// TIA Portal project "XSFW_TIA60401_A3_V14_V15.1" (V15.1) (continued)
   "AuxTempMS050" AT %MW340 : Int;
   "AuxTempMS051" AT %MW342 : Int;
   "AuxTempMS052" AT %MW344 : Int;
   "AuxTempMS053" AT %MW346 : Int;
   "AuxTempMS054" AT %MW348 : Int;
   "AuxTempMS055" AT %MW350 : Int;
   "AuxTempMS056" AT %MW352 : Int;
   "AuxTempMC060" AT %MW354 : Int;
   "AuxTempMC061" AT %MW356 : Int;
   "AuxTempMC062" AT %MW358 : Int;
   "AuxTempMC063" AT %MW360 : Int;
   "AuxTempMC064" AT %MW362 : Int;
   "AuxTempMC065" AT %MW364 : Int;
   "ProxMantBoost1" AT %MD16 : DInt;
   "LimiteMantBoost1" AT %M1.7 : Bool;
   "ProxMantBoost2" AT %MD26 : DInt;
   "LimiteMantBoost2" AT %M2.3 : Bool;
END_VAR

DATA_BLOCK "DB_Fecha"   // DB1
{ S7_Optimized_Access := 'FALSE' }
VERSION : 0.1
   VAR
      STAT0 : Date_And_Time := DT#12-7-5-15:25:53.162;
      STAT1 : Int := 15;
      STAT2 : Int := 25;
      STAT3 : Int := 53;
      STAT4 : Int := 5;
      STAT5 : Int := 7;
      STAT6 : Int := 15;
      STAT7 : Int := 18;
      STAT8 : Int;
      STAT9 : Int := 8;
      STAT10 : Int;
      STAT11 : Word := W#16#15;
      STAT12 : Word := W#16#25;
      STAT13 : Word := W#16#53;
      STAT14 : Word := W#16#5;
      STAT15 : Word := W#16#7;
      STAT16 : Word := W#16#12;
   END_VAR
BEGIN
END_DATA_BLOCK

DATA_BLOCK "Enclavamientos"   // DB28
{ S7_Optimized_Access := 'FALSE' }
VERSION : 0.1
   VAR
      En1 : Bool := true;
      En2 : Bool := true;
      En3 : Bool;
      En4 : Bool;
      En5 : Bool;
      En6 : Bool;
      En7 : Bool;
      En8 : Bool;
      En9 : Bool;
      En10 : Bool;
      En11 : Bool;
      En12 : Bool;
      En13 : Bool;
      En14 : Bool;
      En15 : Bool;
      En16 : Bool;
      En17 : Bool;
      En18 : Bool;
      En19 : Bool;
      En20 : Bool;
      En21 : Bool;
      En22 : Bool;
      En23 : Bool;
      En24 : Bool;
      En25 : Bool;
      En26 : Bool;
      En27 : Bool;
      En28 : Bool;
      En29 : Bool;
      En30 : Bool;
      En31 : Bool;
      En32 : Bool;
      En33 : Bool;
      En34 : Bool;
      En35 : Bool;
      En36 : Bool;
      En37 : Bool;
      En38 : Bool;
      En39 : Bool;
      En40 : Bool;
      En41 : Bool;
      En42 : Bool;
      En43 : Bool;
      En44 : Bool;
      En45 : Bool;
      En46 : Bool;
      En47 : Bool;
      En48 : Bool;
      En49 : Bool;
      En50 : Bool;
      En51 : Bool;
      En52 : Bool;
      En53 : Bool;
      En54 : Bool;
      En55 : Bool;
      En56 : Bool;
      En57 : Bool;
      En58 : Bool;
      En59 : Bool;
      En60 : Bool;
      En61 : Bool;
      En62 : Bool;
      En63 : Bool;
      En64 : Bool;
   END_VAR
BEGIN
END_DATA_BLOCK

// folder: Alarmas

DATA_BLOCK "DB_ALA_PRE"   // DB32
{ S7_Optimized_Access := 'FALSE' }
VERSION : 0.1
   VAR
      x : Bool;   // Ninguna bomba de intercambiador de soplado en marcha
      x1 : Bool;   // Ninguna bomba de chillers de soplado en marcha
      x2 : Bool;   // Ninguna bomba de intercambiador de envasado en marcha
      x3 : Bool;   // Ninguna bomba de chillers de envasado en marcha
      x4 : Bool;   // Ninguna bomba de torre de enfiamiento de chillers en marcha
      x5 : Bool;   // Ningún Chiller de soplado habilitado
      x6 : Bool;   // Ningún chiller de envasado habilitado
      x7 : Bool;   // Alarma Presente en Chiller de soplado Grande
      x8 : Bool;   // Alarma Presente en Chiller de envasado Grande
      x9 : Bool;   // Chiller de soplado Grande en su máxima capacidad
      x10 : Bool;   // Chiller de envasado Grande en su máxima capacidad
      x11 : Bool;   // Falla Térmico MT007
      x12 : Bool;   // Falla Contactor MT007
      x13 : Bool;   // Falla Térmico MT008
      x14 : Bool;   // Falla Contactor MT008
      x15 : Bool;   // Falla Térmico MT009
      x16 : Bool;   // Falla Contactor MT009
      x17 : Bool;   // Falla Térmico MT010
      x18 : Bool;   // Falla Contactor MT010
      x19 : Bool;   // Falla Térmico MP010
      x20 : Bool;   // Falla Contactor MP010
      x21 : Bool;   // Falla Térmico MP011
      x22 : Bool;   // Falla Contactor MP011
      x23 : Bool;   // Falla Térmico MP012
      x24 : Bool;   // Falla Contactor MP012
      x25 : Bool;   // Falla Térmico MP013
      x26 : Bool;   // Falla Contactor MP013
      x27 : Bool;   // Falla Térmico MP018
      x28 : Bool;   // Falla Contactor MP018
      x29 : Bool;   // Falla Térmico MP019
      x30 : Bool;   // Falla Contactor MP019
      x31 : Bool;   // Falla Térmico V001
      x32 : Bool;   // Falla Contactor V001
      x33 : Bool;   // Falla Térmico V002
      x34 : Bool;   // Falla Contactor V002
      x35 : Bool;   // Falla Térmico V003
      x36 : Bool;   // Falla Contactor V003
      x37 : Bool;   // Falla Térmico MC060
      x38 : Bool;   // Falla Contactor MC060
      x39 : Bool;   // Falla Térmico MC061
      x40 : Bool;   // Falla Contactor MC061
      x41 : Bool;   // Falla Térmico MC062
      x42 : Bool;   // Falla Contactor MC062
      x43 : Bool;   // Falla Térmico MC063
      x44 : Bool;   // Falla Contactor MC063
      x45 : Bool;   // Falla Térmico MC064
      x46 : Bool;   // Falla Contactor MC064
      x47 : Bool;   // Falla Térmico MS050
      x48 : Bool;   // Falla Contactor MS050
      x49 : Bool;   // Falla Térmico MS051
      x50 : Bool;   // Falla Contactor MS051
      x51 : Bool;   // Falla Térmico MS052
      x52 : Bool;   // Falla Contactor MS052
      x53 : Bool;   // Falla Térmico MS053
      x54 : Bool;   // Falla Contactor MS053
      x55 : Bool;   // Falla Presostato Chillers
      x56 : Bool;   // Falla Térmico MS054
      x57 : Bool;   // Falla Contactor MS054
      x58 : Bool;   // Falla Térmico MS055
      x59 : Bool;   // Falla Contactor MS055
      x60 : Bool;   // Falla Térmico MV030
      x61 : Bool;   // Falla Contactor MV030
      x62 : Bool;   // Falla Térmico MV031
      x63 : Bool;   // Falla Contactor MV031
      x64 : Bool;   // Falla Térmico MP014
      x65 : Bool;   // Falla Contactor MP014
      x66 : Bool;   // Falla Térmico MP015
      x67 : Bool;   // Falla Contactor MP015
      x68 : Bool;   // Falla Térmico MC001
      x69 : Bool;   // Falla Contactor MC001
      x70 : Bool;   // Falla Térmico MC002
      x71 : Bool;   // Falla Contactor MC002
      x72 : Bool;   // Falla Térmico MC003
      x73 : Bool;   // Falla Contactor MC003
      x74 : Bool;   // Falla Térmico MC004
      x75 : Bool;   // Falla Contactor MC004
      x76 : Bool;   // Falla Térmico MC005
      x77 : Bool;   // Falla Contactor MC005
      x78 : Bool;   // Falla Flujostato Torres Cavaleto
      x79 : Bool;   // Falla Compresor ABC2 Baja Presion de Aceite
      x80 : Bool;   // Falla Compresor ABC2 Baja Presion de Agua
      x81 : Bool;   // Falla Compresor ABC2 Alta Temperatura de Aire
      x82 : Bool;   // Falla Compresor ABC2 Alta Temperatura de agua
      x83 : Bool;   // Falla Compresor ABC3 Baja Presion de Aceite
      x84 : Bool;   // Falla Compresor ABC3 Baja Presion de Agua
      x85 : Bool;   // Falla Compresor ABC3 Alta Temperatura de Aire
      x86 : Bool;   // Falla Compresor ABC3 Alta Temperatura de agua
      x87 : Bool;   // Falla Compresor ABC4 Baja Presion de Aceite
      x88 : Bool;   // Falla Compresor ABC4 Alta Temperatura de Aire
      x89 : Bool;   // Falla Compresor ABC4 Alta Temperatura de Aire
      x90 : Bool;   // Falla Compresor ABC4 Alta Temperatura de agua
      x91 : Bool;   // Falla Compresor ABC5 Baja Presion de Aceite
      x92 : Bool;   // Falla Compresor ABC5 Alta Temperatura de Aire
      x93 : Bool;   // Falla Compresor ABC5 Alta Temperatura de Aire
      x94 : Bool;   // Falla Compresor ABC5 Alta Temperatura de agua
      x95 : Bool;   // Falla Compresor Bellis & MHW28 Baja Presion Aceite
      x96 : Bool;   // Falla Compresor Bellis & MHW28 Baja Presion de Agua
      x97 : Bool;   // Falla Compresor Bellis & MHW28 Alta temperatura de Aire
      x98 : Bool;   // Falla Compresor Bellis & MHW28 Alta temperatura de Agua
      x99 : Bool;   // Falla Compresor Bellis & MHW28 Falla de Flujostato
      x100 : Bool;   // Requiere Marcha MC001
      x101 : Bool;   // Requiere Marcha MC002
      x102 : Bool;   // Requiere Marcha MC003
      x103 : Bool;   // Requiere Marcha MC004
      x104 : Bool;   // Requiere Marcha MC005
      x105 : Bool;   // Falla Conexión con sensor de Temperatura torres de Cavaleto
      x106 : Bool;   // Falla Conexión con sensor de Temperatura torres de Chillers
      x107 : Bool;   // Falla Conexión con sensor de Presión de ALTA
      x108 : Bool;   // Falla Conexión con sensor de Presión de ALTA redundante
      x109 : Bool;   // Falla Conexión con sensor de Presión de Baja
      x110 : Bool;   // Falla Presión de Alta en Límite Mínimo
      x111 : Bool;   // Falla Presión de Alta en demasiado Baja
      x112 : Bool;   // Falla Presión de Alta en demasiado Alta
      x113 : Bool;   // Falla Presión de Alta en Límite Máximo
      x114 : Bool;   // Falla Presión de Baja en Límite Mínimo
      x115 : Bool;   // Falla Presión de Baja en demasiado Baja
      x116 : Bool;   // Falla Presión de Baja en demasiado Alta
      x117 : Bool;   // Falla Presión de Baja en Límite Máximo
      x118 : Bool;   // Falla en chiller de envasado chico
      x119 : Bool;   // Falla en chiller de soplado chico
      x120 : Bool;   // Horas máximas en Compresor 1
      x121 : Bool;   // Horas máximas en Compresor 2
      x122 : Bool;   // Horas máximas en Compresor 3
      x123 : Bool;   // Horas máximas en Compresor 4
      x124 : Bool;   // Horas máximas en Compresor 5
      x125 : Bool;   // Falla algún contactor en Booster
      x126 : Bool;   // Falla algún guardamotor en Booster
      x127 : Bool;   // Presión Alta en Booster
      x128 : Bool;   // Falla algún contactor en Booster 2
      x129 : Bool;   // Falla algún guardamotor en Booster 2
      x130 : Bool;   // Error lectura analógica Presión Boosters
      x131 : Bool;   // Libre
      x132 : Bool;   // Libre
      x133 : Bool;   // Libre
      x134 : Bool;   // Libre
      x135 : Bool;   // Libre
      x136 : Bool;   // Libre
      x137 : Bool;   // Libre
      x138 : Bool;   // Libre
      x139 : Bool;   // Libre
      x140 : Bool;   // Libre
      x141 : Bool;   // Libre
      x142 : Bool;   // Libre
      x143 : Bool;   // Libre
      x144 : Bool;   // ABC1 TTA
      x145 : Bool;   // ABC1TTB
      x146 : Bool;   // ABC1PTA
      x147 : Bool;   // ABC1PTB
      x148 : Bool;   // ABC1Termico
      x149 : Bool;   // ABC1Confirmacion
      x150 : Bool;
      x151 : Bool;
      x152 : Bool;
      x153 : Bool;
      x154 : Bool;
      x155 : Bool;
      x156 : Bool;
      x157 : Bool;
      x158 : Bool;
      x159 : Bool;
      x160 : Bool;
      x161 : Bool;
      x162 : Bool;
      x163 : Bool;
      x164 : Bool;
      x165 : Bool;
      x166 : Bool;
      x167 : Bool;
      x168 : Bool;
      x169 : Bool;
      x170 : Bool;
      x171 : Bool;
      x172 : Bool;
      x173 : Bool;
      x174 : Bool;
      x175 : Bool;
      x176 : Bool;
      x177 : Bool;
      x178 : Bool;
      x179 : Bool;
      x180 : Bool;
      x181 : Bool;
      x182 : Bool;
      x183 : Bool;
      x184 : Bool;
      x185 : Bool;
      x186 : Bool;
      x187 : Bool;
      x188 : Bool;
      x189 : Bool;
      x190 : Bool;
      x191 : Bool;
      x192 : Bool;
      x193 : Bool;
      x194 : Bool;
      x195 : Bool;
      x196 : Bool;
      x197 : Bool;
      x198 : Bool;
      x199 : Bool;
   END_VAR
BEGIN
END_DATA_BLOCK

DATA_BLOCK "DB_ALA_REC"   // DB33
{ S7_Optimized_Access := 'FALSE' }
VERSION : 0.1
   VAR
      x : Bool;   // Ninguna bomba de intercambiador de soplado en marcha
      x1 : Bool;   // Ninguna bomba de chillers de soplado en marcha
      x2 : Bool;   // Ninguna bomba de intercambiador de envasado en marcha
      x3 : Bool;   // Ninguna bomba de chillers de envasado en marcha
      x4 : Bool;   // Ninguna bomba de torre de enfiamiento de chillers en marcha
      x5 : Bool;   // Ningún Chiller de soplado habilitado
      x6 : Bool;   // Ningún chiller de envasado habilitado
      x7 : Bool;   // Alarma Presente en Chiller de soplado Grande
      x8 : Bool;   // Alarma Presente en Chiller de envasado Grande
      x9 : Bool;   // Chiller de soplado Grande en su máxima capacidad
      x10 : Bool;   // Chiller de envasado Grande en su máxima capacidad
      x11 : Bool;   // Falla Térmico MT007
      x12 : Bool;   // Falla Contactor MT007
      x13 : Bool;   // Falla Térmico MT008
      x14 : Bool;   // Falla Contactor MT008
      x15 : Bool;   // Falla Térmico MT009
      x16 : Bool;   // Falla Contactor MT009
      x17 : Bool;   // Falla Térmico MT010
      x18 : Bool;   // Falla Contactor MT010
      x19 : Bool;   // Falla Térmico MP010
      x20 : Bool;   // Falla Contactor MP010
      x21 : Bool;   // Falla Térmico MP011
      x22 : Bool;   // Falla Contactor MP011
      x23 : Bool;   // Falla Térmico MP012
      x24 : Bool;   // Falla Contactor MP012
      x25 : Bool;   // Falla Térmico MP013
      x26 : Bool;   // Falla Contactor MP013
      x27 : Bool;   // Falla Térmico MP018
      x28 : Bool;   // Falla Contactor MP018
      x29 : Bool;   // Falla Térmico MP019
      x30 : Bool;   // Falla Contactor MP019
      x31 : Bool;   // Falla Térmico V001
      x32 : Bool;   // Falla Contactor V001
      x33 : Bool;   // Falla Térmico V002
      x34 : Bool;   // Falla Contactor V002
      x35 : Bool;   // Falla Térmico V003
      x36 : Bool;   // Falla Contactor V003
      x37 : Bool;   // Falla Térmico MC060
      x38 : Bool;   // Falla Contactor MC060
      x39 : Bool;   // Falla Térmico MC061
      x40 : Bool;   // Falla Contactor MC061
      x41 : Bool;   // Falla Térmico MC062
      x42 : Bool;   // Falla Contactor MC062
      x43 : Bool;   // Falla Térmico MC063
      x44 : Bool;   // Falla Contactor MC063
      x45 : Bool;   // Falla Térmico MC064
      x46 : Bool;   // Falla Contactor MC064
      x47 : Bool;   // Falla Térmico MS050
      x48 : Bool;   // Falla Contactor MS050
      x49 : Bool;   // Falla Térmico MS051
      x50 : Bool;   // Falla Contactor MS051
      x51 : Bool;   // Falla Térmico MS052
      x52 : Bool;   // Falla Contactor MS052
      x53 : Bool;   // Falla Térmico MS053
      x54 : Bool;   // Falla Contactor MS053
      x55 : Bool;   // Falla Presostato Chillers
      x56 : Bool;   // Falla Térmico MS054
      x57 : Bool;   // Falla Contactor MS054
      x58 : Bool;   // Falla Térmico MS055
      x59 : Bool;   // Falla Contactor MS055
      x60 : Bool;   // Falla Térmico MV030
      x61 : Bool;   // Falla Contactor MV030
      x62 : Bool;   // Falla Térmico MV031
      x63 : Bool;   // Falla Contactor MV031
      x64 : Bool;   // Falla Térmico MP014
      x65 : Bool;   // Falla Contactor MP014
      x66 : Bool;   // Falla Térmico MP015
      x67 : Bool;   // Falla Contactor MP015
      x68 : Bool;   // Falla Térmico MC001
      x69 : Bool;   // Falla Contactor MC001
      x70 : Bool;   // Falla Térmico MC002
      x71 : Bool;   // Falla Contactor MC002
      x72 : Bool;   // Falla Térmico MC003
      x73 : Bool;   // Falla Contactor MC003
      x74 : Bool;   // Falla Térmico MC004
      x75 : Bool;   // Falla Contactor MC004
      x76 : Bool;   // Falla Térmico MC005
      x77 : Bool;   // Falla Contactor MC005
      x78 : Bool;   // Falla Flujostato Torres Cavaleto
      x79 : Bool;   // Falla Compresor ABC2 Baja Presion de Aceite
      x80 : Bool;   // Falla Compresor ABC2 Baja Presion de Agua
      x81 : Bool;   // Falla Compresor ABC2 Alta Temperatura de Aire
      x82 : Bool;   // Falla Compresor ABC2 Alta Temperatura de agua
      x83 : Bool;   // Falla Compresor ABC3 Baja Presion de Aceite
      x84 : Bool;   // Falla Compresor ABC3 Baja Presion de Agua
      x85 : Bool;   // Falla Compresor ABC3 Alta Temperatura de Aire
      x86 : Bool;   // Falla Compresor ABC3 Alta Temperatura de agua
      x87 : Bool;   // Falla Compresor ABC4 Baja Presion de Aceite
      x88 : Bool;   // Falla Compresor ABC4 Alta Temperatura de Aire
      x89 : Bool;   // Falla Compresor ABC4 Alta Temperatura de Aire
      x90 : Bool;   // Falla Compresor ABC4 Alta Temperatura de agua
      x91 : Bool;   // Falla Compresor ABC5 Baja Presion de Aceite
      x92 : Bool;   // Falla Compresor ABC5 Alta Temperatura de Aire
      x93 : Bool;   // Falla Compresor ABC5 Alta Temperatura de Aire
      x94 : Bool;   // Falla Compresor ABC5 Alta Temperatura de agua
      x95 : Bool;   // Falla Compresor Bellis & MHW28 Baja Presion Aceite
      x96 : Bool;   // Falla Compresor Bellis & MHW28 Baja Presion de Agua
      x97 : Bool;   // Falla Compresor Bellis & MHW28 Alta temperatura de Aire
      x98 : Bool;   // Falla Compresor Bellis & MHW28 Alta temperatura de Agua
      x99 : Bool;   // Falla Compresor Bellis & MHW28 Falla de Flujostato
      x100 : Bool;   // Requiere Marcha MC001
      x101 : Bool;   // Requiere Marcha MC002
      x102 : Bool;   // Requiere Marcha MC003
      x103 : Bool;   // Requiere Marcha MC004
      x104 : Bool;   // Requiere Marcha MC005
      x105 : Bool;   // Falla Conexión con sensor de Temperatura torres de Cavaleto
      x106 : Bool;   // Falla Conexión con sensor de Temperatura torres de Chillers
      x107 : Bool;   // Falla Conexión con sensor de Presión de ALTA
      x108 : Bool;   // Falla Conexión con sensor de Presión de ALTA redundante
      x109 : Bool;   // Falla Conexión con sensor de Presión de Baja
      x110 : Bool;   // Falla Presión de Alta en Límite Mínimo
      x111 : Bool;   // Falla Presión de Alta en demasiado Baja
      x112 : Bool;   // Falla Presión de Alta en demasiado Alta
      x113 : Bool;   // Falla Presión de Alta en Límite Máximo
      x114 : Bool;   // Falla Presión de Baja en Límite Mínimo
      x115 : Bool;   // Falla Presión de Baja en demasiado Baja
      x116 : Bool;   // Falla Presión de Baja en demasiado Alta
      x117 : Bool;   // Falla Presión de Baja en Límite Máximo
      x118 : Bool;   // Falla en chiller de envasado chico
      x119 : Bool;   // Falla en chiller de soplado chico
      x120 : Bool;   // Horas máximas en Compresor 1
      x121 : Bool;   // Horas máximas en Compresor 2
      x122 : Bool;   // Horas máximas en Compresor 3
      x123 : Bool;   // Horas máximas en Compresor 4
      x124 : Bool;   // Horas máximas en Compresor 5
      x125 : Bool;   // Falla algún contactor en Booster
      x126 : Bool;   // Falla algún guardamotor en Booster
      x127 : Bool;   // Presión Alta en Booster
      x128 : Bool;   // Falla algún contactor en Booster 2
      x129 : Bool;   // Falla algún guardamotor en Booster 2
      x130 : Bool;   // Error lectura analógica Presión Boosters
      x131 : Bool;   // Libre
      x132 : Bool;   // Libre
      x133 : Bool;   // Libre
      x134 : Bool;   // Libre
      x135 : Bool;   // Libre
      x136 : Bool;   // Libre
      x137 : Bool;   // Libre
      x138 : Bool;   // Libre
      x139 : Bool;   // Libre
      x140 : Bool;   // Libre
      x141 : Bool;   // Libre
      x142 : Bool;   // Libre
      x143 : Bool;   // Libre
      x144 : Bool;   // ABC1 TTA
      x145 : Bool;   // ABC1TTB
      x146 : Bool;   // ABC1PTA
      x147 : Bool;   // ABC1PTB
      x148 : Bool;   // ABC1Termico
      x149 : Bool;   // ABC1Confirmacion
      x150 : Bool;
      x151 : Bool;
      x152 : Bool;
      x153 : Bool;
      x154 : Bool;
      x155 : Bool;
      x156 : Bool;
      x157 : Bool;
      x158 : Bool;
      x159 : Bool;
      x160 : Bool;
      x161 : Bool;
      x162 : Bool;
      x163 : Bool;
      x164 : Bool;
      x165 : Bool;
      x166 : Bool;
      x167 : Bool;
      x168 : Bool;
      x169 : Bool;
      x170 : Bool;
      x171 : Bool;
      x172 : Bool;
      x173 : Bool;
      x174 : Bool;
      x175 : Bool;
      x176 : Bool;
      x177 : Bool;
      x178 : Bool;
      x179 : Bool;
      x180 : Bool;
      x181 : Bool;
      x182 : Bool;
      x183 : Bool;
      x184 : Bool;
      x185 : Bool;
      x186 : Bool;
      x187 : Bool;
      x188 : Bool;
      x189 : Bool;
      x190 : Bool;
      x191 : Bool;
      x192 : Bool;
      x193 : Bool;
      x194 : Bool;
      x195 : Bool;
      x196 : Bool;
      x197 : Bool;
      x198 : Bool;
      x199 : Bool;
   END_VAR
BEGIN
END_DATA_BLOCK

DATA_BLOCK "DB_ALA_MEM"   // DB34
{ S7_Optimized_Access := 'FALSE' }
VERSION : 0.1
   VAR
      x : Bool;   // Ninguna bomba de intercambiador de soplado en marcha
      x1 : Bool;   // Ninguna bomba de chillers de soplado en marcha
      x2 : Bool;   // Ninguna bomba de intercambiador de envasado en marcha
      x3 : Bool;   // Ninguna bomba de chillers de envasado en marcha
      x4 : Bool;   // Ninguna bomba de torre de enfiamiento de chillers en marcha
      x5 : Bool;   // Ningún Chiller de soplado habilitado
      x6 : Bool;   // Ningún chiller de envasado habilitado
      x7 : Bool;   // Alarma Presente en Chiller de soplado Grande
      x8 : Bool;   // Alarma Presente en Chiller de envasado Grande
      x9 : Bool;   // Chiller de soplado Grande en su máxima capacidad
      x10 : Bool;   // Chiller de envasado Grande en su máxima capacidad
      x11 : Bool;   // Falla Térmico MT007
      x12 : Bool;   // Falla Contactor MT007
      x13 : Bool;   // Falla Térmico MT008
      x14 : Bool;   // Falla Contactor MT008
      x15 : Bool;   // Falla Térmico MT009
      x16 : Bool;   // Falla Contactor MT009
      x17 : Bool;   // Falla Térmico MT010
      x18 : Bool;   // Falla Contactor MT010
      x19 : Bool;   // Falla Térmico MP010
      x20 : Bool;   // Falla Contactor MP010
      x21 : Bool;   // Falla Térmico MP011
      x22 : Bool;   // Falla Contactor MP011
      x23 : Bool;   // Falla Térmico MP012
      x24 : Bool;   // Falla Contactor MP012
      x25 : Bool;   // Falla Térmico MP013
      x26 : Bool;   // Falla Contactor MP013
      x27 : Bool;   // Falla Térmico MP018
      x28 : Bool;   // Falla Contactor MP018
      x29 : Bool;   // Falla Térmico MP019
      x30 : Bool;   // Falla Contactor MP019
      x31 : Bool;   // Falla Térmico V001
      x32 : Bool;   // Falla Contactor V001
      x33 : Bool;   // Falla Térmico V002
      x34 : Bool;   // Falla Contactor V002
      x35 : Bool;   // Falla Térmico V003
      x36 : Bool;   // Falla Contactor V003
      x37 : Bool;   // Falla Térmico MC060
      x38 : Bool;   // Falla Contactor MC060
      x39 : Bool;   // Falla Térmico MC061
      x40 : Bool;   // Falla Contactor MC061
      x41 : Bool;   // Falla Térmico MC062
      x42 : Bool;   // Falla Contactor MC062
      x43 : Bool;   // Falla Térmico MC063
      x44 : Bool;   // Falla Contactor MC063
      x45 : Bool;   // Falla Térmico MC064
      x46 : Bool;   // Falla Contactor MC064
      x47 : Bool;   // Falla Térmico MS050
      x48 : Bool;   // Falla Contactor MS050
      x49 : Bool;   // Falla Térmico MS051
      x50 : Bool;   // Falla Contactor MS051
      x51 : Bool;   // Falla Térmico MS052
      x52 : Bool;   // Falla Contactor MS052
      x53 : Bool;   // Falla Térmico MS053
      x54 : Bool;   // Falla Contactor MS053
      x55 : Bool;   // Falla Presostato Chillers
      x56 : Bool;   // Falla Térmico MS054
      x57 : Bool;   // Falla Contactor MS054
      x58 : Bool;   // Falla Térmico MS055
      x59 : Bool;   // Falla Contactor MS055
      x60 : Bool;   // Falla Térmico MV030
      x61 : Bool;   // Falla Contactor MV030
      x62 : Bool;   // Falla Térmico MV031
      x63 : Bool;   // Falla Contactor MV031
      x64 : Bool;   // Falla Térmico MP014
      x65 : Bool;   // Falla Contactor MP014
      x66 : Bool;   // Falla Térmico MP015
      x67 : Bool;   // Falla Contactor MP015
      x68 : Bool;   // Falla Térmico MC001
      x69 : Bool;   // Falla Contactor MC001
      x70 : Bool;   // Falla Térmico MC002
      x71 : Bool;   // Falla Contactor MC002
      x72 : Bool;   // Falla Térmico MC003
      x73 : Bool;   // Falla Contactor MC003
      x74 : Bool;   // Falla Térmico MC004
      x75 : Bool;   // Falla Contactor MC004
      x76 : Bool;   // Falla Térmico MC005
      x77 : Bool;   // Falla Contactor MC005
      x78 : Bool;   // Falla Flujostato Torres Cavaleto
      x79 : Bool;   // Falla Compresor ABC2 Baja Presion de Aceite
      x80 : Bool;   // Falla Compresor ABC2 Baja Presion de Agua
      x81 : Bool;   // Falla Compresor ABC2 Alta Temperatura de Aire
      x82 : Bool;   // Falla Compresor ABC2 Alta Temperatura de agua
      x83 : Bool;   // Falla Compresor ABC3 Baja Presion de Aceite
      x84 : Bool;   // Falla Compresor ABC3 Baja Presion de Agua
      x85 : Bool;   // Falla Compresor ABC3 Alta Temperatura de Aire
      x86 : Bool;   // Falla Compresor ABC3 Alta Temperatura de agua
      x87 : Bool;   // Falla Compresor ABC4 Baja Presion de Aceite
      x88 : Bool;   // Falla Compresor ABC4 Alta Temperatura de Aire
      x89 : Bool;   // Falla Compresor ABC4 Alta Temperatura de Aire
      x90 : Bool;   // Falla Compresor ABC4 Alta Temperatura de agua
      x91 : Bool;   // Falla Compresor ABC5 Baja Presion de Aceite
      x92 : Bool;   // Falla Compresor ABC5 Alta Temperatura de Aire
      x93 : Bool;   // Falla Compresor ABC5 Alta Temperatura de Aire
      x94 : Bool;   // Falla Compresor ABC5 Alta Temperatura de agua
      x95 : Bool;   // Falla Compresor Bellis & MHW28 Baja Presion Aceite
      x96 : Bool;   // Falla Compresor Bellis & MHW28 Baja Presion de Agua
      x97 : Bool;   // Falla Compresor Bellis & MHW28 Alta temperatura de Aire
      x98 : Bool;   // Falla Compresor Bellis & MHW28 Alta temperatura de Agua
      x99 : Bool;   // Falla Compresor Bellis & MHW28 Falla de Flujostato
      x100 : Bool;   // Requiere Marcha MC001
      x101 : Bool;   // Requiere Marcha MC002
      x102 : Bool;   // Requiere Marcha MC003
      x103 : Bool;   // Requiere Marcha MC004
      x104 : Bool;   // Requiere Marcha MC005
      x105 : Bool;   // Falla Conexión con sensor de Temperatura torres de Cavaleto
      x106 : Bool;   // Falla Conexión con sensor de Temperatura torres de Chillers
      x107 : Bool;   // Falla Conexión con sensor de Presión de ALTA
      x108 : Bool;   // Falla Conexión con sensor de Presión de ALTA redundante
      x109 : Bool;   // Falla Conexión con sensor de Presión de Baja
      x110 : Bool;   // Falla Presión de Alta en Límite Mínimo
      x111 : Bool;   // Falla Presión de Alta en demasiado Baja
      x112 : Bool;   // Falla Presión de Alta en demasiado Alta
      x113 : Bool;   // Falla Presión de Alta en Límite Máximo
      x114 : Bool;   // Falla Presión de Baja en Límite Mínimo
      x115 : Bool;   // Falla Presión de Baja en demasiado Baja
      x116 : Bool;   // Falla Presión de Baja en demasiado Alta
      x117 : Bool;   // Falla Presión de Baja en Límite Máximo
      x118 : Bool;   // Falla en chiller de envasado chico
      x119 : Bool;   // Falla en chiller de soplado chico
      x120 : Bool;   // Horas máximas en Compresor 1
      x121 : Bool;   // Horas máximas en Compresor 2
      x122 : Bool;   // Horas máximas en Compresor 3
      x123 : Bool;   // Horas máximas en Compresor 4
      x124 : Bool;   // Horas máximas en Compresor 5
      x125 : Bool;   // Falla algún contactor en Booster
      x126 : Bool;   // Falla algún guardamotor en Booster
      x127 : Bool;   // Presión Alta en Booster
      x128 : Bool;   // Falla algún contactor en Booster 2
      x129 : Bool;   // Falla algún guardamotor en Booster 2
      x130 : Bool;   // Error lectura analógica Presión Boosters
      x131 : Bool;   // Libre
      x132 : Bool;   // Libre
      x133 : Bool;   // Libre
      x134 : Bool;   // Libre
      x135 : Bool;   // Libre
      x136 : Bool;   // Libre
      x137 : Bool;   // Libre
      x138 : Bool;   // Libre
      x139 : Bool;   // Libre
      x140 : Bool;   // Libre
      x141 : Bool;   // Libre
      x142 : Bool;   // Libre
      x143 : Bool;   // Libre
      x144 : Bool;   // ABC1 TTA
      x145 : Bool;   // ABC1TTB
      x146 : Bool;   // ABC1PTA
      x147 : Bool;   // ABC1PTB
      x148 : Bool;   // ABC1Termico
      x149 : Bool;   // ABC1Confirmacion
      x150 : Bool;
      x151 : Bool;
      x152 : Bool;
      x153 : Bool;
      x154 : Bool;
      x155 : Bool;
      x156 : Bool;
      x157 : Bool;
      x158 : Bool;
      x159 : Bool;
      x160 : Bool;
      x161 : Bool;
      x162 : Bool;
      x163 : Bool;
      x164 : Bool;
      x165 : Bool;
      x166 : Bool;
      x167 : Bool;
      x168 : Bool;
      x169 : Bool;
      x170 : Bool;
      x171 : Bool;
      x172 : Bool;
      x173 : Bool;
      x174 : Bool;
      x175 : Bool;
      x176 : Bool;
      x177 : Bool;
      x178 : Bool;
      x179 : Bool;
      x180 : Bool;
      x181 : Bool;
      x182 : Bool;
      x183 : Bool;
      x184 : Bool;
      x185 : Bool;
      x186 : Bool;
      x187 : Bool;
      x188 : Bool;
      x189 : Bool;
      x190 : Bool;
      x191 : Bool;
      x192 : Bool;
      x193 : Bool;
      x194 : Bool;
      x195 : Bool;
      x196 : Bool;
      x197 : Bool;
      x198 : Bool;
      x199 : Bool;
   END_VAR
BEGIN
END_DATA_BLOCK

DATA_BLOCK "DB_COM_REC"   // DB35
{ S7_Optimized_Access := 'FALSE' }
VERSION : 0.1
   VAR
      x : Bool;   // Ninguna bomba de intercambiador de soplado en marcha
      x1 : Bool;   // Ninguna bomba de chillers de soplado en marcha
      x2 : Bool;   // Ninguna bomba de intercambiador de envasado en marcha
      x3 : Bool;   // Ninguna bomba de chillers de envasado en marcha
      x4 : Bool;   // Ninguna bomba de torre de enfiamiento de chillers en marcha
      x5 : Bool;   // Ningún Chiller de soplado habilitado
      x6 : Bool;   // Ningún chiller de envasado habilitado
      x7 : Bool;   // Alarma Presente en Chiller de soplado Grande
      x8 : Bool;   // Alarma Presente en Chiller de envasado Grande
      x9 : Bool;   // Chiller de soplado Grande en su máxima capacidad
      x10 : Bool;   // Chiller de envasado Grande en su máxima capacidad
      x11 : Bool;   // Falla Térmico MT007
      x12 : Bool;   // Falla Contactor MT007
      x13 : Bool;   // Falla Térmico MT008
      x14 : Bool;   // Falla Contactor MT008
      x15 : Bool;   // Falla Térmico MT009
      x16 : Bool;   // Falla Contactor MT009
      x17 : Bool;   // Falla Térmico MT010
      x18 : Bool;   // Falla Contactor MT010
      x19 : Bool;   // Falla Térmico MP010
      x20 : Bool;   // Falla Contactor MP010
      x21 : Bool;   // Falla Térmico MP011
      x22 : Bool;   // Falla Contactor MP011
      x23 : Bool;   // Falla Térmico MP012
      x24 : Bool;   // Falla Contactor MP012
      x25 : Bool;   // Falla Térmico MP013
      x26 : Bool;   // Falla Contactor MP013
      x27 : Bool;   // Falla Térmico MP018
      x28 : Bool;   // Falla Contactor MP018
      x29 : Bool;   // Falla Térmico MP019
      x30 : Bool;   // Falla Contactor MP019
      x31 : Bool;   // Falla Térmico V001
      x32 : Bool;   // Falla Contactor V001
      x33 : Bool;   // Falla Térmico V002
      x34 : Bool;   // Falla Contactor V002
      x35 : Bool;   // Falla Térmico V003
      x36 : Bool;   // Falla Contactor V003
      x37 : Bool;   // Falla Térmico MC060
      x38 : Bool;   // Falla Contactor MC060
      x39 : Bool;   // Falla Térmico MC061
      x40 : Bool;   // Falla Contactor MC061
      x41 : Bool;   // Falla Térmico MC062
      x42 : Bool;   // Falla Contactor MC062
      x43 : Bool;   // Falla Térmico MC063
      x44 : Bool;   // Falla Contactor MC063
      x45 : Bool;   // Falla Térmico MC064
      x46 : Bool;   // Falla Contactor MC064
      x47 : Bool;   // Falla Térmico MS050
      x48 : Bool;   // Falla Contactor MS050
      x49 : Bool;   // Falla Térmico MS051
      x50 : Bool;   // Falla Contactor MS051
      x51 : Bool;   // Falla Térmico MS052
      x52 : Bool;   // Falla Contactor MS052
      x53 : Bool;   // Falla Térmico MS053
      x54 : Bool;   // Falla Contactor MS053
      x55 : Bool;   // Falla Presostato Chillers
      x56 : Bool;   // Falla Térmico MS054
      x57 : Bool;   // Falla Contactor MS054
      x58 : Bool;   // Falla Térmico MS055
      x59 : Bool;   // Falla Contactor MS055
      x60 : Bool;   // Falla Térmico MV030
      x61 : Bool;   // Falla Contactor MV030
      x62 : Bool;   // Falla Térmico MV031
      x63 : Bool;   // Falla Contactor MV031
      x64 : Bool;   // Falla Térmico MP014
      x65 : Bool;   // Falla Contactor MP014
      x66 : Bool;   // Falla Térmico MP015
      x67 : Bool;   // Falla Contactor MP015
      x68 : Bool;   // Falla Térmico MC001
      x69 : Bool;   // Falla Contactor MC001
      x70 : Bool;   // Falla Térmico MC002
      x71 : Bool;   // Falla Contactor MC002
      x72 : Bool;   // Falla Térmico MC003
      x73 : Bool;   // Falla Contactor MC003
      x74 : Bool;   // Falla Térmico MC004
      x75 : Bool;   // Falla Contactor MC004
      x76 : Bool;   // Falla Térmico MC005
      x77 : Bool;   // Falla Contactor MC005
      x78 : Bool;   // Falla Flujostato Torres Cavaleto
      x79 : Bool;   // Falla Compresor ABC2 Baja Presion de Aceite
      x80 : Bool;   // Falla Compresor ABC2 Baja Presion de Agua
      x81 : Bool;   // Falla Compresor ABC2 Alta Temperatura de Aire
      x82 : Bool;   // Falla Compresor ABC2 Alta Temperatura de agua
      x83 : Bool;   // Falla Compresor ABC3 Baja Presion de Aceite
      x84 : Bool;   // Falla Compresor ABC3 Baja Presion de Agua
      x85 : Bool;   // Falla Compresor ABC3 Alta Temperatura de Aire
      x86 : Bool;   // Falla Compresor ABC3 Alta Temperatura de agua
      x87 : Bool;   // Falla Compresor ABC4 Baja Presion de Aceite
      x88 : Bool;   // Falla Compresor ABC4 Alta Temperatura de Aire
      x89 : Bool;   // Falla Compresor ABC4 Alta Temperatura de Aire
      x90 : Bool;   // Falla Compresor ABC4 Alta Temperatura de agua
      x91 : Bool;   // Falla Compresor ABC5 Baja Presion de Aceite
      x92 : Bool;   // Falla Compresor ABC5 Alta Temperatura de Aire
      x93 : Bool;   // Falla Compresor ABC5 Alta Temperatura de Aire
      x94 : Bool;   // Falla Compresor ABC5 Alta Temperatura de agua
      x95 : Bool;   // Falla Compresor Bellis & MHW28 Baja Presion Aceite
      x96 : Bool;   // Falla Compresor Bellis & MHW28 Baja Presion de Agua
      x97 : Bool;   // Falla Compresor Bellis & MHW28 Alta temperatura de Aire
      x98 : Bool;   // Falla Compresor Bellis & MHW28 Alta temperatura de Agua
      x99 : Bool;   // Falla Compresor Bellis & MHW28 Falla de Flujostato
      x100 : Bool;   // Requiere Marcha MC001
      x101 : Bool;   // Requiere Marcha MC002
      x102 : Bool;   // Requiere Marcha MC003
      x103 : Bool;   // Requiere Marcha MC004
      x104 : Bool;   // Requiere Marcha MC005
      x105 : Bool;   // Falla Conexión con sensor de Temperatura torres de Cavaleto
      x106 : Bool;   // Falla Conexión con sensor de Temperatura torres de Chillers
      x107 : Bool;   // Falla Conexión con sensor de Presión de ALTA
      x108 : Bool;   // Falla Conexión con sensor de Presión de ALTA redundante
      x109 : Bool;   // Falla Conexión con sensor de Presión de Baja
      x110 : Bool;   // Falla Presión de Alta en Límite Mínimo
      x111 : Bool;   // Falla Presión de Alta en demasiado Baja
      x112 : Bool;   // Falla Presión de Alta en demasiado Alta
      x113 : Bool;   // Falla Presión de Alta en Límite Máximo
      x114 : Bool;   // Falla Presión de Baja en Límite Mínimo
      x115 : Bool;   // Falla Presión de Baja en demasiado Baja
      x116 : Bool;   // Falla Presión de Baja en demasiado Alta
      x117 : Bool;   // Falla Presión de Baja en Límite Máximo
      x118 : Bool;   // Falla en chiller de envasado chico
      x119 : Bool;   // Falla en chiller de soplado chico
      x120 : Bool;   // Horas máximas en Compresor 1
      x121 : Bool;   // Horas máximas en Compresor 2
      x122 : Bool;   // Horas máximas en Compresor 3
      x123 : Bool;   // Horas máximas en Compresor 4
      x124 : Bool;   // Horas máximas en Compresor 5
      x125 : Bool;   // Falla algún contactor en Booster
      x126 : Bool;   // Falla algún guardamotor en Booster
      x127 : Bool;   // Presión Alta en Booster
      x128 : Bool;   // Falla algún contactor en Booster 2
      x129 : Bool;   // Falla algún guardamotor en Booster 2
      x130 : Bool;   // Error lectura analógica Presión Boosters
      x131 : Bool;   // Libre
      x132 : Bool;   // Libre
      x133 : Bool;   // Libre
      x134 : Bool;   // Libre
      x135 : Bool;   // Libre
      x136 : Bool;   // Libre
      x137 : Bool;   // Libre
      x138 : Bool;   // Libre
      x139 : Bool;   // Libre
      x140 : Bool;   // Libre
      x141 : Bool;   // Libre
      x142 : Bool;   // Libre
      x143 : Bool;   // Libre
      x144 : Bool;
      x145 : Bool;
      x146 : Bool;
      x147 : Bool;
      x148 : Bool;
      x149 : Bool;
      x150 : Bool;
      x151 : Bool;
      x152 : Bool;
      x153 : Bool;
      x154 : Bool;
      x155 : Bool;
      x156 : Bool;
      x157 : Bool;
      x158 : Bool;
      x159 : Bool;
      x160 : Bool;
      x161 : Bool;
      x162 : Bool;
      x163 : Bool;
      x164 : Bool;
      x165 : Bool;
      x166 : Bool;
      x167 : Bool;
      x168 : Bool;
      x169 : Bool;
      x170 : Bool;
      x171 : Bool;
      x172 : Bool;
      x173 : Bool;
      x174 : Bool;
      x175 : Bool;
      x176 : Bool;
      x177 : Bool;
      x178 : Bool;
      x179 : Bool;
      x180 : Bool;
      x181 : Bool;
      x182 : Bool;
      x183 : Bool;
      x184 : Bool;
      x185 : Bool;
      x186 : Bool;
      x187 : Bool;
      x188 : Bool;
      x189 : Bool;
      x190 : Bool;
      x191 : Bool;
      x192 : Bool;
      x193 : Bool;
      x194 : Bool;
      x195 : Bool;
      x196 : Bool;
      x197 : Bool;
      x198 : Bool;
      x199 : Bool;
   END_VAR
BEGIN
END_DATA_BLOCK

DATA_BLOCK "DB_COM__REC_FLANCO"   // DB36
{ S7_Optimized_Access := 'FALSE' }
VERSION : 0.1
   VAR
      x : Bool;   // Ninguna bomba de intercambiador de soplado en marcha
      x1 : Bool;   // Ninguna bomba de chillers de soplado en marcha
      x2 : Bool;   // Ninguna bomba de intercambiador de envasado en marcha
      x3 : Bool;   // Ninguna bomba de chillers de envasado en marcha
      x4 : Bool;   // Ninguna bomba de torre de enfiamiento de chillers en marcha
      x5 : Bool;   // Ningún Chiller de soplado habilitado
      x6 : Bool;   // Ningún chiller de envasado habilitado
      x7 : Bool;   // Alarma Presente en Chiller de soplado Grande
      x8 : Bool;   // Alarma Presente en Chiller de envasado Grande
      x9 : Bool;   // Chiller de soplado Grande en su máxima capacidad
      x10 : Bool;   // Chiller de envasado Grande en su máxima capacidad
      x11 : Bool;   // Falla Térmico MT007
      x12 : Bool;   // Falla Contactor MT007
      x13 : Bool;   // Falla Térmico MT008
      x14 : Bool;   // Falla Contactor MT008
      x15 : Bool;   // Falla Térmico MT009
      x16 : Bool;   // Falla Contactor MT009
      x17 : Bool;   // Falla Térmico MT010
      x18 : Bool;   // Falla Contactor MT010
      x19 : Bool;   // Falla Térmico MP010
      x20 : Bool;   // Falla Contactor MP010
      x21 : Bool;   // Falla Térmico MP011
      x22 : Bool;   // Falla Contactor MP011
      x23 : Bool;   // Falla Térmico MP012
      x24 : Bool;   // Falla Contactor MP012
      x25 : Bool;   // Falla Térmico MP013
      x26 : Bool;   // Falla Contactor MP013
      x27 : Bool;   // Falla Térmico MP018
      x28 : Bool;   // Falla Contactor MP018
      x29 : Bool;   // Falla Térmico MP019
      x30 : Bool;   // Falla Contactor MP019
      x31 : Bool;   // Falla Térmico V001
      x32 : Bool;   // Falla Contactor V001
      x33 : Bool;   // Falla Térmico V002
      x34 : Bool;   // Falla Contactor V002
      x35 : Bool;   // Falla Térmico V003
      x36 : Bool;   // Falla Contactor V003
      x37 : Bool;   // Falla Térmico MC060
      x38 : Bool;   // Falla Contactor MC060
      x39 : Bool;   // Falla Térmico MC061
      x40 : Bool;   // Falla Contactor MC061
      x41 : Bool;   // Falla Térmico MC062
      x42 : Bool;   // Falla Contactor MC062
      x43 : Bool;   // Falla Térmico MC063
      x44 : Bool;   // Falla Contactor MC063
      x45 : Bool;   // Falla Térmico MC064
      x46 : Bool;   // Falla Contactor MC064
      x47 : Bool;   // Falla Térmico MS050
      x48 : Bool;   // Falla Contactor MS050
      x49 : Bool;   // Falla Térmico MS051
      x50 : Bool;   // Falla Contactor MS051
      x51 : Bool;   // Falla Térmico MS052
      x52 : Bool;   // Falla Contactor MS052
      x53 : Bool;   // Falla Térmico MS053
      x54 : Bool;   // Falla Contactor MS053
      x55 : Bool;   // Falla Presostato Chillers
      x56 : Bool;   // Falla Térmico MS054
      x57 : Bool;   // Falla Contactor MS054
      x58 : Bool;   // Falla Térmico MS055
      x59 : Bool;   // Falla Contactor MS055
      x60 : Bool;   // Falla Térmico MV030
      x61 : Bool;   // Falla Contactor MV030
      x62 : Bool;   // Falla Térmico MV031
      x63 : Bool;   // Falla Contactor MV031
      x64 : Bool;   // Falla Térmico MP014
      x65 : Bool;   // Falla Contactor MP014
      x66 : Bool;   // Falla Térmico MP015
      x67 : Bool;   // Falla Contactor MP015
      x68 : Bool;   // Falla Térmico MC001
      x69 : Bool;   // Falla Contactor MC001
      x70 : Bool;   // Falla Térmico MC002
      x71 : Bool;   // Falla Contactor MC002
      x72 : Bool;   // Falla Térmico MC003
      x73 : Bool;   // Falla Contactor MC003
      x74 : Bool;   // Falla Térmico MC004
      x75 : Bool;   // Falla Contactor MC004
      x76 : Bool;   // Falla Térmico MC005
      x77 : Bool;   // Falla Contactor MC005
      x78 : Bool;   // Falla Flujostato Torres Cavaleto
      x79 : Bool;   // Falla Compresor ABC2 Baja Presion de Aceite
      x80 : Bool;   // Falla Compresor ABC2 Baja Presion de Agua
      x81 : Bool;   // Falla Compresor ABC2 Alta Temperatura de Aire
      x82 : Bool;   // Falla Compresor ABC2 Alta Temperatura de agua
      x83 : Bool;   // Falla Compresor ABC3 Baja Presion de Aceite
      x84 : Bool;   // Falla Compresor ABC3 Baja Presion de Agua
      x85 : Bool;   // Falla Compresor ABC3 Alta Temperatura de Aire
      x86 : Bool;   // Falla Compresor ABC3 Alta Temperatura de agua
      x87 : Bool;   // Falla Compresor ABC4 Baja Presion de Aceite
      x88 : Bool;   // Falla Compresor ABC4 Alta Temperatura de Aire
      x89 : Bool;   // Falla Compresor ABC4 Alta Temperatura de Aire
      x90 : Bool;   // Falla Compresor ABC4 Alta Temperatura de agua
      x91 : Bool;   // Falla Compresor ABC5 Baja Presion de Aceite
      x92 : Bool;   // Falla Compresor ABC5 Alta Temperatura de Aire
      x93 : Bool;   // Falla Compresor ABC5 Alta Temperatura de Aire
      x94 : Bool;   // Falla Compresor ABC5 Alta Temperatura de agua
      x95 : Bool;   // Falla Compresor Bellis & MHW28 Baja Presion Aceite
      x96 : Bool;   // Falla Compresor Bellis & MHW28 Baja Presion de Agua
      x97 : Bool;   // Falla Compresor Bellis & MHW28 Alta temperatura de Aire
      x98 : Bool;   // Falla Compresor Bellis & MHW28 Alta temperatura de Agua
      x99 : Bool;   // Falla Compresor Bellis & MHW28 Falla de Flujostato
      x100 : Bool;   // Requiere Marcha MC001
      x101 : Bool;   // Requiere Marcha MC002
      x102 : Bool;   // Requiere Marcha MC003
      x103 : Bool;   // Requiere Marcha MC004
      x104 : Bool;   // Requiere Marcha MC005
      x105 : Bool;   // Falla Conexión con sensor de Temperatura torres de Cavaleto
      x106 : Bool;   // Falla Conexión con sensor de Temperatura torres de Chillers
      x107 : Bool;   // Falla Conexión con sensor de Presión de ALTA
      x108 : Bool;   // Falla Conexión con sensor de Presión de ALTA redundante
      x109 : Bool;   // Falla Conexión con sensor de Presión de Baja
      x110 : Bool;   // Falla Presión de Alta en Límite Mínimo
      x111 : Bool;   // Falla Presión de Alta en demasiado Baja
      x112 : Bool;   // Falla Presión de Alta en demasiado Alta
      x113 : Bool;   // Falla Presión de Alta en Límite Máximo
      x114 : Bool;   // Falla Presión de Baja en Límite Mínimo
      x115 : Bool;   // Falla Presión de Baja en demasiado Baja
      x116 : Bool;   // Falla Presión de Baja en demasiado Alta
      x117 : Bool;   // Falla Presión de Baja en Límite Máximo
      x118 : Bool;   // Falla en chiller de envasado chico
      x119 : Bool;   // Falla en chiller de soplado chico
      x120 : Bool;   // Horas máximas en Compresor 1
      x121 : Bool;   // Horas máximas en Compresor 2
      x122 : Bool;   // Horas máximas en Compresor 3
      x123 : Bool;   // Horas máximas en Compresor 4
      x124 : Bool;   // Horas máximas en Compresor 5
      x125 : Bool;   // Falla algún contactor en Booster
      x126 : Bool;   // Falla algún guardamotor en Booster
      x127 : Bool;   // Presión Alta en Booster
      x128 : Bool;   // Falla algún contactor en Booster 2
      x129 : Bool;   // Falla algún guardamotor en Booster 2
      x130 : Bool;   // Error lectura analógica Presión Boosters
      x131 : Bool;   // Libre
      x132 : Bool;   // Libre
      x133 : Bool;   // Libre
      x134 : Bool;   // Libre
      x135 : Bool;   // Libre
      x136 : Bool;   // Libre
      x137 : Bool;   // Libre
      x138 : Bool;   // Libre
      x139 : Bool;   // Libre
      x140 : Bool;   // Libre
      x141 : Bool;   // Libre
      x142 : Bool;   // Libre
      x143 : Bool;   // Libre
      x144 : Bool;
      x145 : Bool;
      x146 : Bool;
      x147 : Bool;
      x148 : Bool;
      x149 : Bool;
      x150 : Bool;
      x151 : Bool;
      x152 : Bool;
      x153 : Bool;
      x154 : Bool;
      x155 : Bool;
      x156 : Bool;
      x157 : Bool;
      x158 : Bool;
      x159 : Bool;
      x160 : Bool;
      x161 : Bool;
      x162 : Bool;
      x163 : Bool;
      x164 : Bool;
      x165 : Bool;
      x166 : Bool;
      x167 : Bool;
      x168 : Bool;
      x169 : Bool;
      x170 : Bool;
      x171 : Bool;
      x172 : Bool;
      x173 : Bool;
      x174 : Bool;
      x175 : Bool;
      x176 : Bool;
      x177 : Bool;
      x178 : Bool;
      x179 : Bool;
      x180 : Bool;
      x181 : Bool;
      x182 : Bool;
      x183 : Bool;
      x184 : Bool;
      x185 : Bool;
      x186 : Bool;
      x187 : Bool;
      x188 : Bool;
      x189 : Bool;
      x190 : Bool;
      x191 : Bool;
      x192 : Bool;
      x193 : Bool;
      x194 : Bool;
      x195 : Bool;
      x196 : Bool;
      x197 : Bool;
      x198 : Bool;
      x199 : Bool;
   END_VAR
BEGIN
END_DATA_BLOCK

